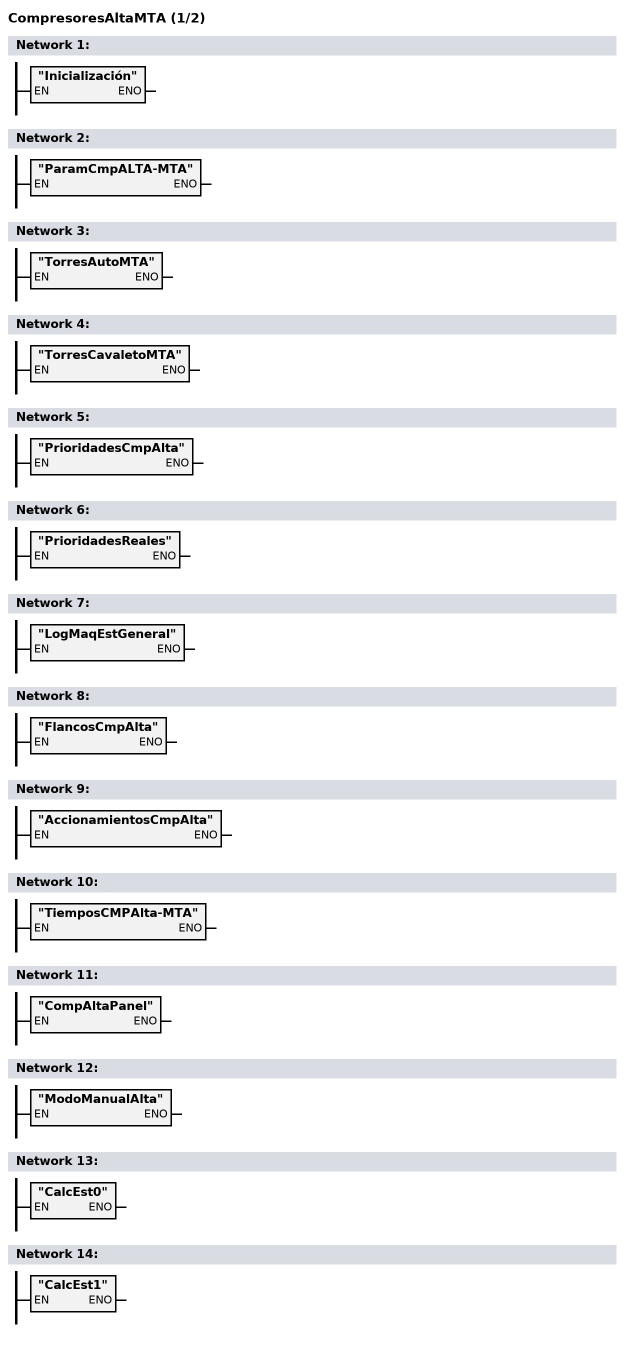
   RUNG wire#powerrail
      "Inicialización"()
   END_RUNG
   // the same network as SCL:
   "Inicialización"();
END_REGION

REGION Network 2
   RUNG wire#powerrail
      "ParamCmpALTA-MTA"()
   END_RUNG
   // the same network as SCL:
   "ParamCmpALTA-MTA"();
END_REGION

REGION Network 3
   RUNG wire#powerrail
      "TorresAutoMTA"()
   END_RUNG
   // the same network as SCL:
   "TorresAutoMTA"();
END_REGION

REGION Network 4
   RUNG wire#powerrail
      "TorresCavaletoMTA"()
   END_RUNG
   // the same network as SCL:
   "TorresCavaletoMTA"();
END_REGION

REGION Network 5
   RUNG wire#powerrail
      "PrioridadesCmpAlta"()
   END_RUNG
   // the same network as SCL:
   "PrioridadesCmpAlta"();
END_REGION

REGION Network 6
   RUNG wire#powerrail
      "PrioridadesReales"()
   END_RUNG
   // the same network as SCL:
   "PrioridadesReales"();
END_REGION

REGION Network 7
   RUNG wire#powerrail
      "LogMaqEstGeneral"()
   END_RUNG
   // the same network as SCL:
   "LogMaqEstGeneral"();
END_REGION

REGION Network 8
   RUNG wire#powerrail
      "FlancosCmpAlta"()
   END_RUNG
   // the same network as SCL:
   "FlancosCmpAlta"();
END_REGION

REGION Network 9
   RUNG wire#powerrail
      "AccionamientosCmpAlta"()
   END_RUNG
   // the same network as SCL:
   "AccionamientosCmpAlta"();
END_REGION

REGION Network 10
   RUNG wire#powerrail
      "TiemposCMPAlta-MTA"()
   END_RUNG
   // the same network as SCL:
   "TiemposCMPAlta-MTA"();
END_REGION

REGION Network 11
   RUNG wire#powerrail
      "CompAltaPanel"()
   END_RUNG
   // the same network as SCL:
   "CompAltaPanel"();
END_REGION

REGION Network 12
   RUNG wire#powerrail
      "ModoManualAlta"()
   END_RUNG
   // the same network as SCL:
   "ModoManualAlta"();
END_REGION

REGION Network 13
   RUNG wire#powerrail
      "CalcEst0"()
   END_RUNG
   // the same network as SCL:
   "CalcEst0"();
END_REGION

REGION Network 14
   RUNG wire#powerrail
      "CalcEst1"()
   END_RUNG
   // the same network as SCL:
   "CalcEst1"();
END_REGION

REGION Network 15
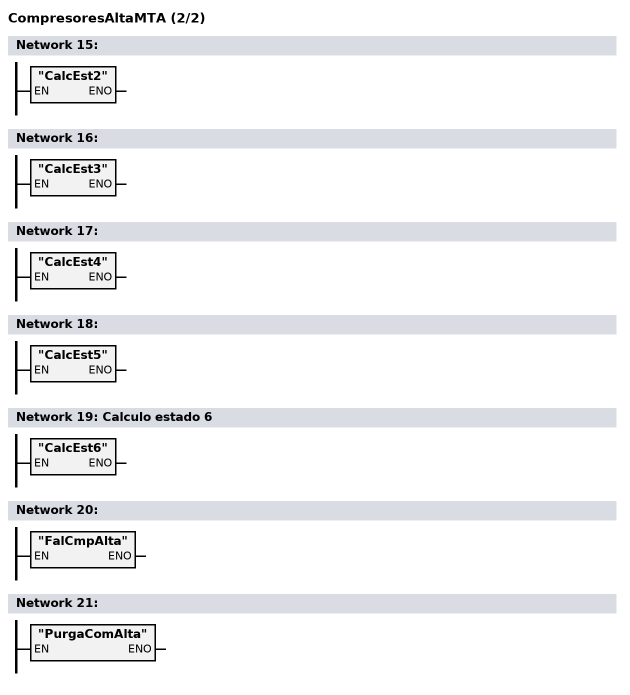
   RUNG wire#powerrail
      "CalcEst2"()
   END_RUNG
   // the same network as SCL:
   "CalcEst2"();
END_REGION

REGION Network 16
   RUNG wire#powerrail
      "CalcEst3"()
   END_RUNG
   // the same network as SCL:
   "CalcEst3"();
END_REGION

REGION Network 17
   RUNG wire#powerrail
      "CalcEst4"()
   END_RUNG
   // the same network as SCL:
   "CalcEst4"();
END_REGION

REGION Network 18
   RUNG wire#powerrail
      "CalcEst5"()
   END_RUNG
   // the same network as SCL:
   "CalcEst5"();
END_REGION

REGION Network 19: Calculo estado 6
   RUNG wire#powerrail
      "CalcEst6"()
   END_RUNG
   // the same network as SCL:
   "CalcEst6"();
END_REGION

REGION Network 20
   RUNG wire#powerrail
      "FalCmpAlta"()
   END_RUNG
   // the same network as SCL:
   "FalCmpAlta"();
END_REGION

REGION Network 21
   RUNG wire#powerrail
      "PurgaComAlta"()
   END_RUNG
   // the same network as SCL:
   "PurgaComAlta"();
END_REGION
END_FUNCTION

FUNCTION "ParamCmpALTA-MTA" : Void   // FC30, LAD
{ S7_Optimized_Access := 'FALSE' }
VERSION : 0.1
BEGIN

REGION Network 1
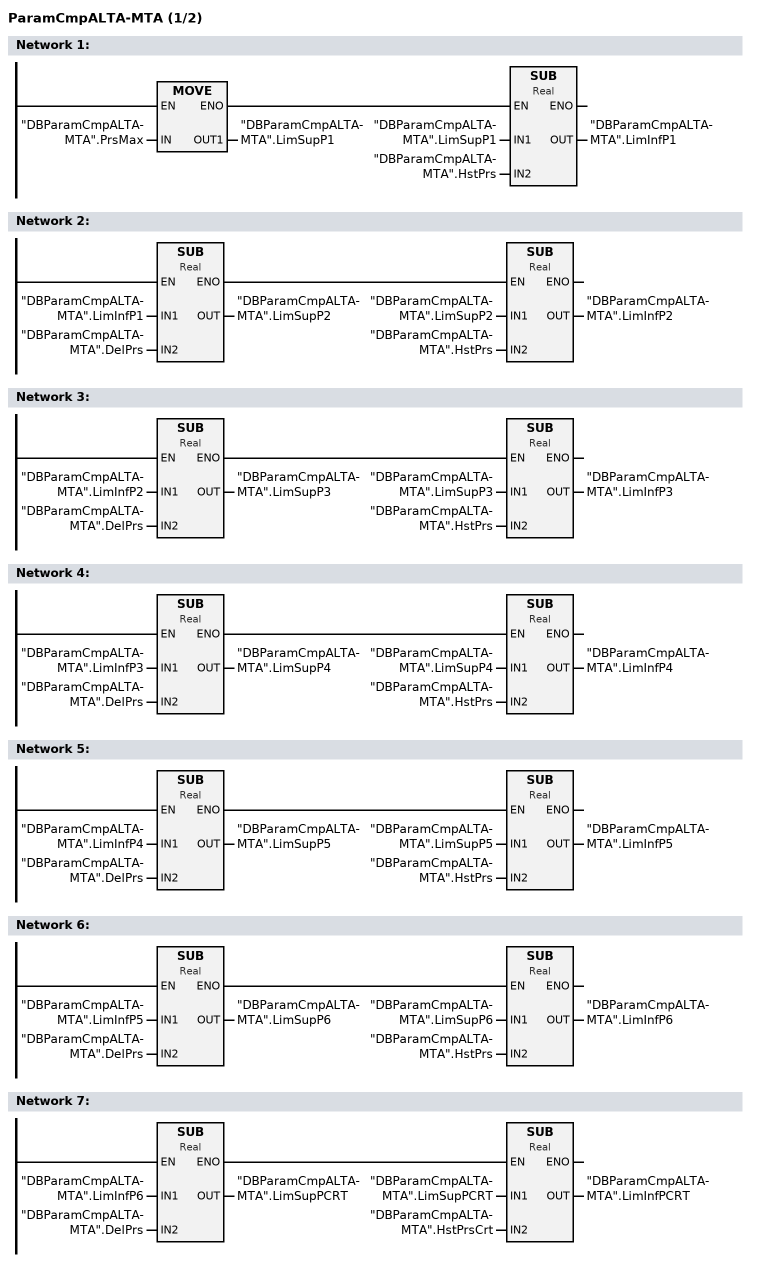
   RUNG wire#powerrail
      { S7_GenerateENO := "TRUE" } Move(in := "DBParamCmpALTA-MTA".PrsMax, out1 => "DBParamCmpALTA-MTA".LimSupP1)
      { S7_Templates := "SrcType := Real"; S7_GenerateENO := "TRUE" } Sub(in1 := "DBParamCmpALTA-MTA".LimSupP1, in2 := "DBParamCmpALTA-MTA".HstPrs, out => "DBParamCmpALTA-MTA".LimInfP1)
   END_RUNG
   // the same network as SCL:
   // ENO of a box is taken as its EN; it also drops when the box reports an error
   "DBParamCmpALTA-MTA".LimSupP1 := "DBParamCmpALTA-MTA".PrsMax;
   "DBParamCmpALTA-MTA".LimInfP1 := "DBParamCmpALTA-MTA".LimSupP1 - "DBParamCmpALTA-MTA".HstPrs;
END_REGION

REGION Network 2
   RUNG wire#powerrail
      { S7_Templates := "SrcType := Real"; S7_GenerateENO := "TRUE" } Sub(in1 := "DBParamCmpALTA-MTA".LimInfP1, in2 := "DBParamCmpALTA-MTA".DelPrs, out => "DBParamCmpALTA-MTA".LimSupP2)
      { S7_Templates := "SrcType := Real"; S7_GenerateENO := "TRUE" } Sub(in1 := "DBParamCmpALTA-MTA".LimSupP2, in2 := "DBParamCmpALTA-MTA".HstPrs, out => "DBParamCmpALTA-MTA".LimInfP2)
   END_RUNG
   // the same network as SCL:
   // ENO of a box is taken as its EN; it also drops when the box reports an error
   "DBParamCmpALTA-MTA".LimSupP2 := "DBParamCmpALTA-MTA".LimInfP1 - "DBParamCmpALTA-MTA".DelPrs;
   "DBParamCmpALTA-MTA".LimInfP2 := "DBParamCmpALTA-MTA".LimSupP2 - "DBParamCmpALTA-MTA".HstPrs;
END_REGION

REGION Network 3
   RUNG wire#powerrail
      { S7_Templates := "SrcType := Real"; S7_GenerateENO := "TRUE" } Sub(in1 := "DBParamCmpALTA-MTA".LimInfP2, in2 := "DBParamCmpALTA-MTA".DelPrs, out => "DBParamCmpALTA-MTA".LimSupP3)
      { S7_Templates := "SrcType := Real"; S7_GenerateENO := "TRUE" } Sub(in1 := "DBParamCmpALTA-MTA".LimSupP3, in2 := "DBParamCmpALTA-MTA".HstPrs, out => "DBParamCmpALTA-MTA".LimInfP3)
   END_RUNG
   // the same network as SCL:
   // ENO of a box is taken as its EN; it also drops when the box reports an error
   "DBParamCmpALTA-MTA".LimSupP3 := "DBParamCmpALTA-MTA".LimInfP2 - "DBParamCmpALTA-MTA".DelPrs;
   "DBParamCmpALTA-MTA".LimInfP3 := "DBParamCmpALTA-MTA".LimSupP3 - "DBParamCmpALTA-MTA".HstPrs;
END_REGION

REGION Network 4
   RUNG wire#powerrail
      { S7_Templates := "SrcType := Real"; S7_GenerateENO := "TRUE" } Sub(in1 := "DBParamCmpALTA-MTA".LimInfP3, in2 := "DBParamCmpALTA-MTA".DelPrs, out => "DBParamCmpALTA-MTA".LimSupP4)
      { S7_Templates := "SrcType := Real"; S7_GenerateENO := "TRUE" } Sub(in1 := "DBParamCmpALTA-MTA".LimSupP4, in2 := "DBParamCmpALTA-MTA".HstPrs, out => "DBParamCmpALTA-MTA".LimInfP4)
   END_RUNG
   // the same network as SCL:
   // ENO of a box is taken as its EN; it also drops when the box reports an error
   "DBParamCmpALTA-MTA".LimSupP4 := "DBParamCmpALTA-MTA".LimInfP3 - "DBParamCmpALTA-MTA".DelPrs;
   "DBParamCmpALTA-MTA".LimInfP4 := "DBParamCmpALTA-MTA".LimSupP4 - "DBParamCmpALTA-MTA".HstPrs;
END_REGION

REGION Network 5
   RUNG wire#powerrail
      { S7_Templates := "SrcType := Real"; S7_GenerateENO := "TRUE" } Sub(in1 := "DBParamCmpALTA-MTA".LimInfP4, in2 := "DBParamCmpALTA-MTA".DelPrs, out => "DBParamCmpALTA-MTA".LimSupP5)
      { S7_Templates := "SrcType := Real"; S7_GenerateENO := "TRUE" } Sub(in1 := "DBParamCmpALTA-MTA".LimSupP5, in2 := "DBParamCmpALTA-MTA".HstPrs, out => "DBParamCmpALTA-MTA".LimInfP5)
   END_RUNG
   // the same network as SCL:
   // ENO of a box is taken as its EN; it also drops when the box reports an error
   "DBParamCmpALTA-MTA".LimSupP5 := "DBParamCmpALTA-MTA".LimInfP4 - "DBParamCmpALTA-MTA".DelPrs;
   "DBParamCmpALTA-MTA".LimInfP5 := "DBParamCmpALTA-MTA".LimSupP5 - "DBParamCmpALTA-MTA".HstPrs;
END_REGION

REGION Network 6
   RUNG wire#powerrail
      { S7_Templates := "SrcType := Real"; S7_GenerateENO := "TRUE" } Sub(in1 := "DBParamCmpALTA-MTA".LimInfP5, in2 := "DBParamCmpALTA-MTA".DelPrs, out => "DBParamCmpALTA-MTA".LimSupP6)
      { S7_Templates := "SrcType := Real"; S7_GenerateENO := "TRUE" } Sub(in1 := "DBParamCmpALTA-MTA".LimSupP6, in2 := "DBParamCmpALTA-MTA".HstPrs, out => "DBParamCmpALTA-MTA".LimInfP6)
   END_RUNG
   // the same network as SCL:
   // ENO of a box is taken as its EN; it also drops when the box reports an error
   "DBParamCmpALTA-MTA".LimSupP6 := "DBParamCmpALTA-MTA".LimInfP5 - "DBParamCmpALTA-MTA".DelPrs;
   "DBParamCmpALTA-MTA".LimInfP6 := "DBParamCmpALTA-MTA".LimSupP6 - "DBParamCmpALTA-MTA".HstPrs;
END_REGION

REGION Network 7
   RUNG wire#powerrail
      { S7_Templates := "SrcType := Real"; S7_GenerateENO := "TRUE" } Sub(in1 := "DBParamCmpALTA-MTA".LimInfP6, in2 := "DBParamCmpALTA-MTA".DelPrs, out => "DBParamCmpALTA-MTA".LimSupPCRT)
      { S7_Templates := "SrcType := Real"; S7_GenerateENO := "TRUE" } Sub(in1 := "DBParamCmpALTA-MTA".LimSupPCRT, in2 := "DBParamCmpALTA-MTA".HstPrsCrt, out => "DBParamCmpALTA-MTA".LimInfPCRT)
   END_RUNG
   // the same network as SCL:
   // ENO of a box is taken as its EN; it also drops when the box reports an error
   "DBParamCmpALTA-MTA".LimSupPCRT := "DBParamCmpALTA-MTA".LimInfP6 - "DBParamCmpALTA-MTA".DelPrs;
   "DBParamCmpALTA-MTA".LimInfPCRT := "DBParamCmpALTA-MTA".LimSupPCRT - "DBParamCmpALTA-MTA".HstPrsCrt;
END_REGION

REGION Network 8: Falla General Flujostato Cavaleto
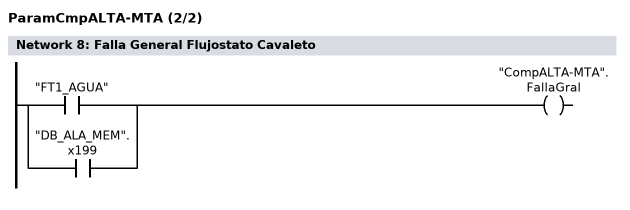
   RUNG wire#powerrail
      Contact( "FT1_AGUA" )
      wire#w1
      Coil( "CompALTA-MTA".FallaGral )
   END_RUNG
   RUNG wire#powerrail
      Contact( "DB_ALA_MEM".x199 )
   END_RUNG wire#w1
   // the same network as SCL:
   "CompALTA-MTA".FallaGral := "FT1_AGUA" OR "DB_ALA_MEM".x199;
END_REGION
END_FUNCTION

FUNCTION "TiemposCMPAlta-MTA" : Void   // FC31, LAD
{ S7_Optimized_Access := 'FALSE' }
VERSION : 0.1
   VAR_TEMP
      TEMP0 : Int;
   END_VAR
   VAR_TEMP   // added for the SCL form of the ladder/FBD networks
      _s5time1 : S5Time;
   END_VAR
BEGIN

REGION Network 1
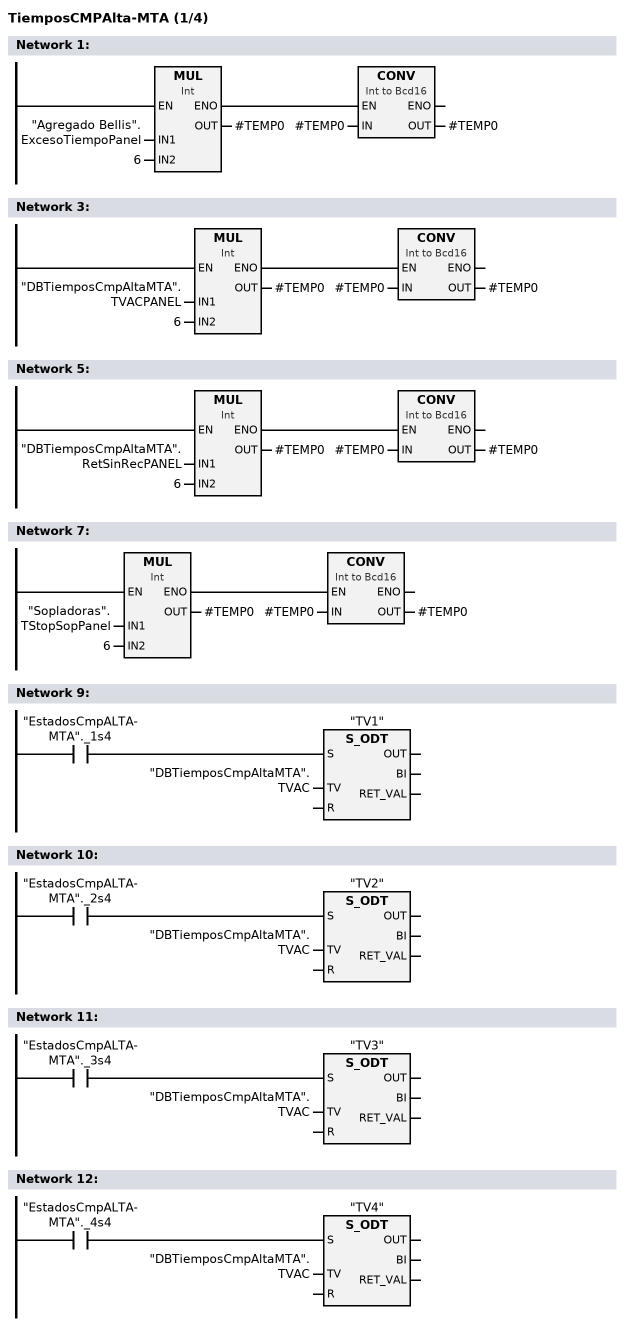
   RUNG wire#powerrail
      { S7_Templates := "SrcType := Int"; S7_GenerateENO := "TRUE" } Mul(in1 := "Agregado Bellis".ExcesoTiempoPanel, in2 := 6, out => #TEMP0)
      { S7_Templates := "[SrcType := Int, DestType := Bcd16]"; S7_GenerateENO := "TRUE" } Convert(in := #TEMP0, out => #TEMP0)
   END_RUNG
   // the same network as SCL:
   // ENO of a box is taken as its EN; it also drops when the box reports an error
   #TEMP0 := "Agregado Bellis".ExcesoTiempoPanel * 6;
   #TEMP0 := INT_TO_BCD16(#TEMP0);
END_REGION

REGION Network 2 (STL)
         L     12288;
         L     #TEMP0;
         OW;
         T     "Agregado Bellis".ExcesoTiempo;
         NOP   0;
END_REGION

REGION Network 3
   RUNG wire#powerrail
      { S7_Templates := "SrcType := Int"; S7_GenerateENO := "TRUE" } Mul(in1 := "DBTiemposCmpAltaMTA".TVACPANEL, in2 := 6, out => #TEMP0)
      { S7_Templates := "[SrcType := Int, DestType := Bcd16]"; S7_GenerateENO := "TRUE" } Convert(in := #TEMP0, out => #TEMP0)
   END_RUNG
   // the same network as SCL:
   // ENO of a box is taken as its EN; it also drops when the box reports an error
   #TEMP0 := "DBTiemposCmpAltaMTA".TVACPANEL * 6;
   #TEMP0 := INT_TO_BCD16(#TEMP0);
END_REGION

REGION Network 4 (STL)
         L     12288;
         L     #TEMP0;
         OW;
         T     "DBTiemposCmpAltaMTA".TVAC;
         NOP   0;
END_REGION

REGION Network 5
   RUNG wire#powerrail
      { S7_Templates := "SrcType := Int"; S7_GenerateENO := "TRUE" } Mul(in1 := "DBTiemposCmpAltaMTA".RetSinRecPANEL, in2 := 6, out => #TEMP0)
      { S7_Templates := "[SrcType := Int, DestType := Bcd16]"; S7_GenerateENO := "TRUE" } Convert(in := #TEMP0, out => #TEMP0)
   END_RUNG
   // the same network as SCL:
   // ENO of a box is taken as its EN; it also drops when the box reports an error
   #TEMP0 := "DBTiemposCmpAltaMTA".RetSinRecPANEL * 6;
   #TEMP0 := INT_TO_BCD16(#TEMP0);
END_REGION

REGION Network 6 (STL)
         L     12288;
         L     #TEMP0;
         OW;
         T     "DBTiemposCmpAltaMTA".RetSinRec;
         NOP   0;
END_REGION

REGION Network 7
   RUNG wire#powerrail
      { S7_Templates := "SrcType := Int"; S7_GenerateENO := "TRUE" } Mul(in1 := "Sopladoras".TStopSopPanel, in2 := 6, out => #TEMP0)
      { S7_Templates := "[SrcType := Int, DestType := Bcd16]"; S7_GenerateENO := "TRUE" } Convert(in := #TEMP0, out => #TEMP0)
   END_RUNG
   // the same network as SCL:
   // ENO of a box is taken as its EN; it also drops when the box reports an error
   #TEMP0 := "Sopladoras".TStopSopPanel * 6;
   #TEMP0 := INT_TO_BCD16(#TEMP0);
END_REGION

REGION Network 8 (STL)
         L     12288;
         L     #TEMP0;
         OW;
         T     "Sopladoras".TStopSop;
         NOP   0;
END_REGION

REGION Network 9
   RUNG wire#powerrail
      Contact( "EstadosCmpALTA-MTA"._1s4 )
      S_ODT(T_NO := "TV1", TV := "DBTiemposCmpAltaMTA".TVAC, R :=, BI =>, RET_VAL =>)
   END_RUNG
   // the same network as SCL:
   #_s5time1 := S_ODT(T_NO := "TV1", S := "EstadosCmpALTA-MTA"._1s4, TV := "DBTiemposCmpAltaMTA".TVAC);
END_REGION

REGION Network 10
   RUNG wire#powerrail
      Contact( "EstadosCmpALTA-MTA"._2s4 )
      S_ODT(T_NO := "TV2", TV := "DBTiemposCmpAltaMTA".TVAC, R :=, BI =>, RET_VAL =>)
   END_RUNG
   // the same network as SCL:
   #_s5time1 := S_ODT(T_NO := "TV2", S := "EstadosCmpALTA-MTA"._2s4, TV := "DBTiemposCmpAltaMTA".TVAC);
END_REGION

REGION Network 11
   RUNG wire#powerrail
      Contact( "EstadosCmpALTA-MTA"._3s4 )
      S_ODT(T_NO := "TV3", TV := "DBTiemposCmpAltaMTA".TVAC, R :=, BI =>, RET_VAL =>)
   END_RUNG
   // the same network as SCL:
   #_s5time1 := S_ODT(T_NO := "TV3", S := "EstadosCmpALTA-MTA"._3s4, TV := "DBTiemposCmpAltaMTA".TVAC);
END_REGION

REGION Network 12
   RUNG wire#powerrail
      Contact( "EstadosCmpALTA-MTA"._4s4 )
      S_ODT(T_NO := "TV4", TV := "DBTiemposCmpAltaMTA".TVAC, R :=, BI =>, RET_VAL =>)
   END_RUNG
   // the same network as SCL:
   #_s5time1 := S_ODT(T_NO := "TV4", S := "EstadosCmpALTA-MTA"._4s4, TV := "DBTiemposCmpAltaMTA".TVAC);
END_REGION

REGION Network 13
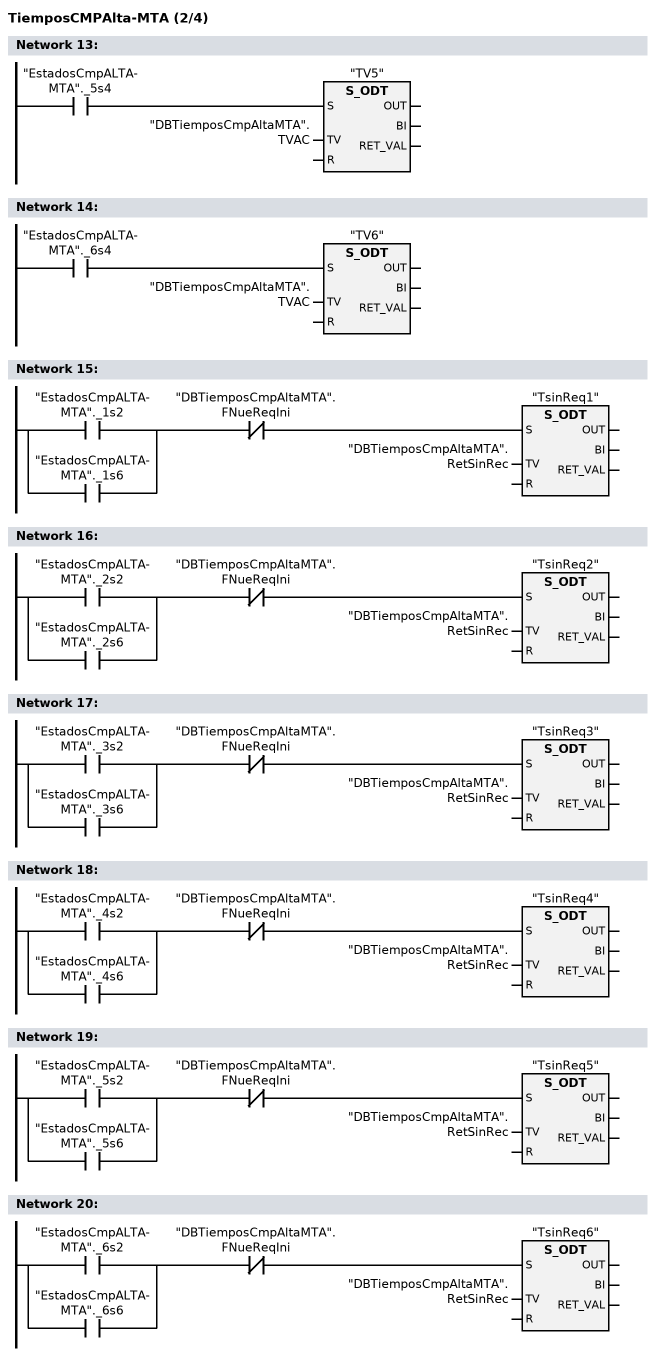
   RUNG wire#powerrail
      Contact( "EstadosCmpALTA-MTA"._5s4 )
      S_ODT(T_NO := "TV5", TV := "DBTiemposCmpAltaMTA".TVAC, R :=, BI =>, RET_VAL =>)
   END_RUNG
   // the same network as SCL:
   #_s5time1 := S_ODT(T_NO := "TV5", S := "EstadosCmpALTA-MTA"._5s4, TV := "DBTiemposCmpAltaMTA".TVAC);
END_REGION

REGION Network 14
   RUNG wire#powerrail
      Contact( "EstadosCmpALTA-MTA"._6s4 )
      S_ODT(T_NO := "TV6", TV := "DBTiemposCmpAltaMTA".TVAC, R :=, BI =>, RET_VAL =>)
   END_RUNG
   // the same network as SCL:
   #_s5time1 := S_ODT(T_NO := "TV6", S := "EstadosCmpALTA-MTA"._6s4, TV := "DBTiemposCmpAltaMTA".TVAC);
END_REGION

REGION Network 15
   RUNG wire#powerrail
      Contact( "EstadosCmpALTA-MTA"._1s2 )
      wire#w1
      I_Contact( "DBTiemposCmpAltaMTA".FNueReqIni )
      S_ODT(T_NO := "TsinReq1", TV := "DBTiemposCmpAltaMTA".RetSinRec, R :=, BI =>, RET_VAL =>)
   END_RUNG
   RUNG wire#powerrail
      Contact( "EstadosCmpALTA-MTA"._1s6 )
   END_RUNG wire#w1
   // the same network as SCL:
   #_s5time1 := S_ODT(T_NO := "TsinReq1",
                      S := ("EstadosCmpALTA-MTA"._1s2 OR "EstadosCmpALTA-MTA"._1s6) AND NOT "DBTiemposCmpAltaMTA".FNueReqIni,
                      TV := "DBTiemposCmpAltaMTA".RetSinRec);
END_REGION

REGION Network 16
   RUNG wire#powerrail
      Contact( "EstadosCmpALTA-MTA"._2s2 )
      wire#w1
      I_Contact( "DBTiemposCmpAltaMTA".FNueReqIni )
      S_ODT(T_NO := "TsinReq2", TV := "DBTiemposCmpAltaMTA".RetSinRec, R :=, BI =>, RET_VAL =>)
   END_RUNG
   RUNG wire#powerrail
      Contact( "EstadosCmpALTA-MTA"._2s6 )
   END_RUNG wire#w1
   // the same network as SCL:
   #_s5time1 := S_ODT(T_NO := "TsinReq2",
                      S := ("EstadosCmpALTA-MTA"._2s2 OR "EstadosCmpALTA-MTA"._2s6) AND NOT "DBTiemposCmpAltaMTA".FNueReqIni,
                      TV := "DBTiemposCmpAltaMTA".RetSinRec);
END_REGION

REGION Network 17
   RUNG wire#powerrail
      Contact( "EstadosCmpALTA-MTA"._3s2 )
      wire#w1
      I_Contact( "DBTiemposCmpAltaMTA".FNueReqIni )
      S_ODT(T_NO := "TsinReq3", TV := "DBTiemposCmpAltaMTA".RetSinRec, R :=, BI =>, RET_VAL =>)
   END_RUNG
   RUNG wire#powerrail
      Contact( "EstadosCmpALTA-MTA"._3s6 )
   END_RUNG wire#w1
   // the same network as SCL:
   #_s5time1 := S_ODT(T_NO := "TsinReq3",
                      S := ("EstadosCmpALTA-MTA"._3s2 OR "EstadosCmpALTA-MTA"._3s6) AND NOT "DBTiemposCmpAltaMTA".FNueReqIni,
                      TV := "DBTiemposCmpAltaMTA".RetSinRec);
END_REGION

REGION Network 18
   RUNG wire#powerrail
      Contact( "EstadosCmpALTA-MTA"._4s2 )
      wire#w1
      I_Contact( "DBTiemposCmpAltaMTA".FNueReqIni )
      S_ODT(T_NO := "TsinReq4", TV := "DBTiemposCmpAltaMTA".RetSinRec, R :=, BI =>, RET_VAL =>)
   END_RUNG
   RUNG wire#powerrail
      Contact( "EstadosCmpALTA-MTA"._4s6 )
   END_RUNG wire#w1
   // the same network as SCL:
   #_s5time1 := S_ODT(T_NO := "TsinReq4",
                      S := ("EstadosCmpALTA-MTA"._4s2 OR "EstadosCmpALTA-MTA"._4s6) AND NOT "DBTiemposCmpAltaMTA".FNueReqIni,
                      TV := "DBTiemposCmpAltaMTA".RetSinRec);
END_REGION

REGION Network 19
   RUNG wire#powerrail
      Contact( "EstadosCmpALTA-MTA"._5s2 )
      wire#w1
      I_Contact( "DBTiemposCmpAltaMTA".FNueReqIni )
      S_ODT(T_NO := "TsinReq5", TV := "DBTiemposCmpAltaMTA".RetSinRec, R :=, BI =>, RET_VAL =>)
   END_RUNG
   RUNG wire#powerrail
      Contact( "EstadosCmpALTA-MTA"._5s6 )
   END_RUNG wire#w1
   // the same network as SCL:
   #_s5time1 := S_ODT(T_NO := "TsinReq5",
                      S := ("EstadosCmpALTA-MTA"._5s2 OR "EstadosCmpALTA-MTA"._5s6) AND NOT "DBTiemposCmpAltaMTA".FNueReqIni,
                      TV := "DBTiemposCmpAltaMTA".RetSinRec);
END_REGION

REGION Network 20
   RUNG wire#powerrail
      Contact( "EstadosCmpALTA-MTA"._6s2 )
      wire#w1
      I_Contact( "DBTiemposCmpAltaMTA".FNueReqIni )
      S_ODT(T_NO := "TsinReq6", TV := "DBTiemposCmpAltaMTA".RetSinRec, R :=, BI =>, RET_VAL =>)
   END_RUNG
   RUNG wire#powerrail
      Contact( "EstadosCmpALTA-MTA"._6s6 )
   END_RUNG wire#w1
   // the same network as SCL:
   #_s5time1 := S_ODT(T_NO := "TsinReq6",
                      S := ("EstadosCmpALTA-MTA"._6s2 OR "EstadosCmpALTA-MTA"._6s6) AND NOT "DBTiemposCmpAltaMTA".FNueReqIni,
                      TV := "DBTiemposCmpAltaMTA".RetSinRec);
END_REGION

REGION Network 21
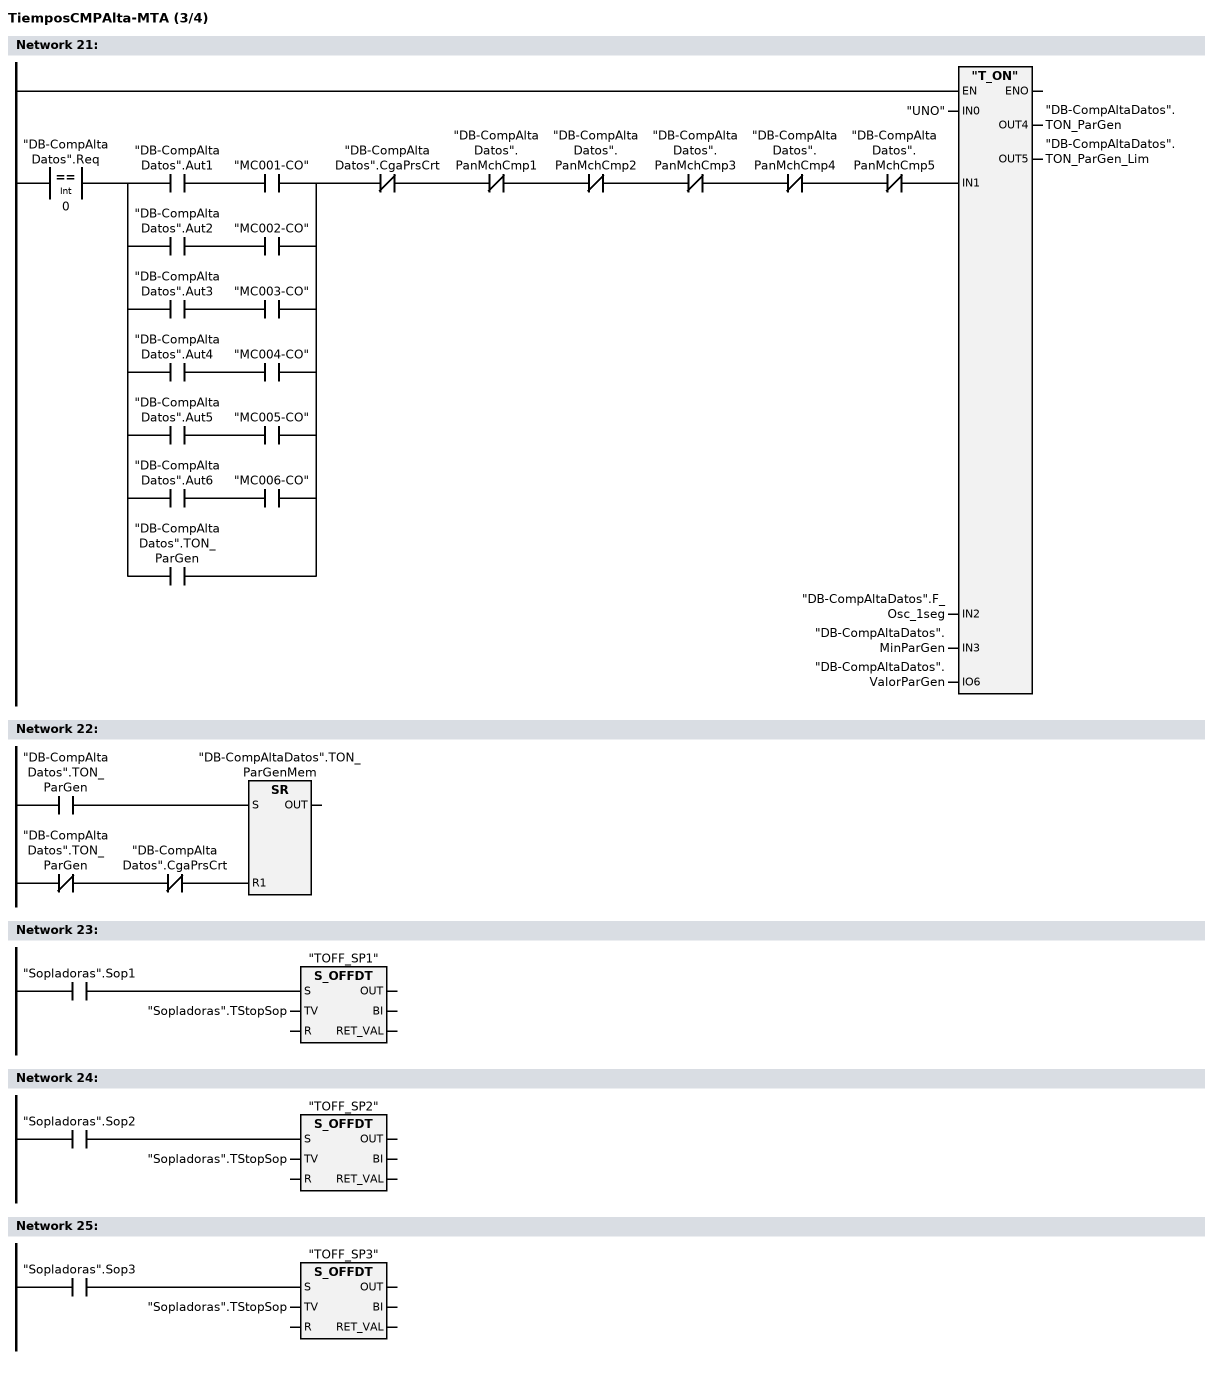
   RUNG wire#powerrail
      "T_ON"(IN1 := wire#w3, IN0 := "UNO", IN2 := "DB-CompAltaDatos".F_Osc_1seg, IN3 := "DB-CompAltaDatos".MinParGen, IO6 := "DB-CompAltaDatos".ValorParGen, OUT4 => "DB-CompAltaDatos".TON_ParGen, OUT5 => "DB-CompAltaDatos".TON_ParGen_Lim)
   END_RUNG
   RUNG wire#powerrail
      { S7_Templates := "SrcType := Int" } EQ_Contact(in1 := "DB-CompAltaDatos".Req, in2 := 0)
      wire#w1
      Contact( "DB-CompAltaDatos".Aut1 )
      Contact( "MC001-CO" )
      wire#w2
      I_Contact( "DB-CompAltaDatos".CgaPrsCrt )
      I_Contact( "DB-CompAltaDatos".PanMchCmp1 )
      I_Contact( "DB-CompAltaDatos".PanMchCmp2 )
      I_Contact( "DB-CompAltaDatos".PanMchCmp3 )
      I_Contact( "DB-CompAltaDatos".PanMchCmp4 )
      I_Contact( "DB-CompAltaDatos".PanMchCmp5 )
   END_RUNG wire#w3
   RUNG wire#w1
      Contact( "DB-CompAltaDatos".Aut2 )
      Contact( "MC002-CO" )
   END_RUNG wire#w2
   RUNG wire#w1
      Contact( "DB-CompAltaDatos".Aut3 )
      Contact( "MC003-CO" )
   END_RUNG wire#w2
   RUNG wire#w1
      Contact( "DB-CompAltaDatos".Aut4 )
      Contact( "MC004-CO" )
   END_RUNG wire#w2
   RUNG wire#w1
      Contact( "DB-CompAltaDatos".Aut5 )
      Contact( "MC005-CO" )
   END_RUNG wire#w2
   RUNG wire#w1
      Contact( "DB-CompAltaDatos".Aut6 )
      Contact( "MC006-CO" )
   END_RUNG wire#w2
   RUNG wire#w1
      Contact( "DB-CompAltaDatos".TON_ParGen )
   END_RUNG wire#w2
   // the same network as SCL:
   "T_ON"(IN0 := "UNO",
          IN1 := ("DB-CompAltaDatos".Req = 0) AND (("DB-CompAltaDatos".Aut1 AND "MC001-CO") OR ("DB-CompAltaDatos".Aut2 AND "MC002-CO") OR ("DB-CompAltaDatos".Aut3 AND "MC003-CO") OR ("DB-CompAltaDatos".Aut4 AND "MC004-CO") OR ("DB-CompAltaDatos".Aut5 AND "MC005-CO") OR ("DB-CompAltaDatos".Aut6 AND "MC006-CO") OR "DB-CompAltaDatos".TON_ParGen) AND NOT "DB-CompAltaDatos".CgaPrsCrt AND NOT "DB-CompAltaDatos".PanMchCmp1 AND NOT "DB-CompAltaDatos".PanMchCmp2 AND NOT "DB-CompAltaDatos".PanMchCmp3 AND NOT "DB-CompAltaDatos".PanMchCmp4 AND NOT "DB-CompAltaDatos".PanMchCmp5,
          IN2 := "DB-CompAltaDatos".F_Osc_1seg,
          IN3 := "DB-CompAltaDatos".MinParGen,
          IO6 := "DB-CompAltaDatos".ValorParGen,
          OUT4 => "DB-CompAltaDatos".TON_ParGen,
          OUT5 => "DB-CompAltaDatos".TON_ParGen_Lim);
END_REGION

REGION Network 22
   RUNG wire#powerrail
      Contact( "DB-CompAltaDatos".TON_ParGen )
      S_SR(operand := "DB-CompAltaDatos".TON_ParGenMem, r1 := wire#w1)
   END_RUNG
   RUNG wire#powerrail
      I_Contact( "DB-CompAltaDatos".TON_ParGen )
      I_Contact( "DB-CompAltaDatos".CgaPrsCrt )
   END_RUNG wire#w1
   // the same network as SCL:
   IF "DB-CompAltaDatos".TON_ParGen THEN
       "DB-CompAltaDatos".TON_ParGenMem := TRUE;   // SR flip-flop
   END_IF;
   IF NOT "DB-CompAltaDatos".TON_ParGen AND NOT "DB-CompAltaDatos".CgaPrsCrt THEN
       "DB-CompAltaDatos".TON_ParGenMem := FALSE;
   END_IF;
END_REGION

REGION Network 23
   RUNG wire#powerrail
      Contact( "Sopladoras".Sop1 )
      S_OFFDT(T_NO := "TOFF_SP1", TV := "Sopladoras".TStopSop, R :=, BI =>, RET_VAL =>)
   END_RUNG
   // the same network as SCL:
   #_s5time1 := S_OFFDT(T_NO := "TOFF_SP1", TV := "Sopladoras".TStopSop, S := "Sopladoras".Sop1);
END_REGION

REGION Network 24
   RUNG wire#powerrail
      Contact( "Sopladoras".Sop2 )
      S_OFFDT(T_NO := "TOFF_SP2", TV := "Sopladoras".TStopSop, R :=, BI =>, RET_VAL =>)
   END_RUNG
   // the same network as SCL:
   #_s5time1 := S_OFFDT(T_NO := "TOFF_SP2", TV := "Sopladoras".TStopSop, S := "Sopladoras".Sop2);
END_REGION

REGION Network 25
   RUNG wire#powerrail
      Contact( "Sopladoras".Sop3 )
      S_OFFDT(T_NO := "TOFF_SP3", TV := "Sopladoras".TStopSop, R :=, BI =>, RET_VAL =>)
   END_RUNG
   // the same network as SCL:
   #_s5time1 := S_OFFDT(T_NO := "TOFF_SP3", TV := "Sopladoras".TStopSop, S := "Sopladoras".Sop3);
END_REGION

REGION Network 26
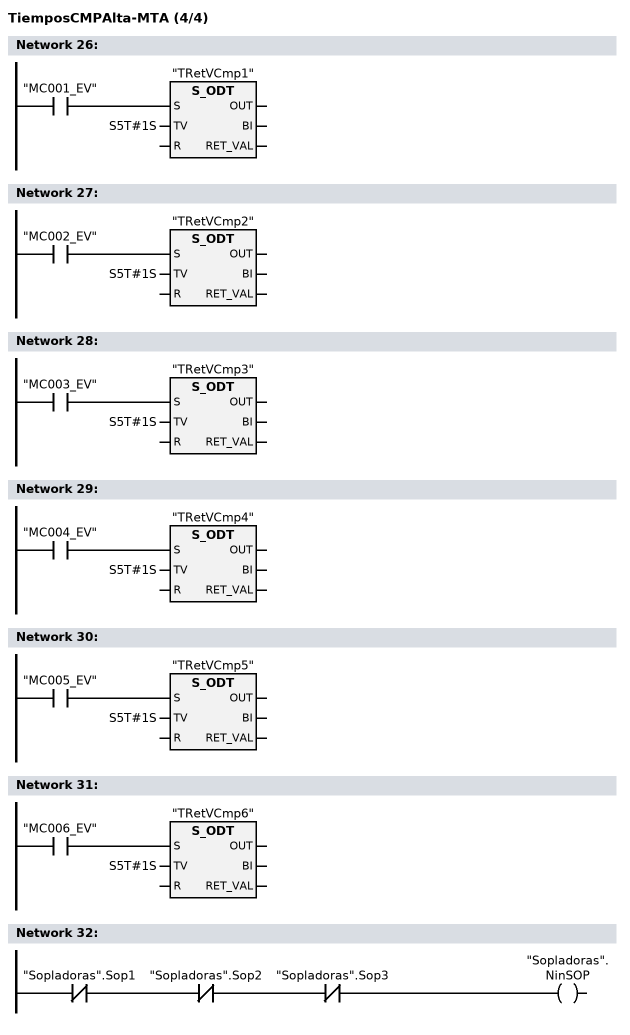
   RUNG wire#powerrail
      Contact( "MC001_EV" )
      S_ODT(T_NO := "TRetVCmp1", TV := S5T#1S, R :=, BI =>, RET_VAL =>)
   END_RUNG
   // the same network as SCL:
   #_s5time1 := S_ODT(T_NO := "TRetVCmp1", TV := S5T#1S, S := "MC001_EV");
END_REGION

REGION Network 27
   RUNG wire#powerrail
      Contact( "MC002_EV" )
      S_ODT(T_NO := "TRetVCmp2", TV := S5T#1S, R :=, BI =>, RET_VAL =>)
   END_RUNG
   // the same network as SCL:
   #_s5time1 := S_ODT(T_NO := "TRetVCmp2", TV := S5T#1S, S := "MC002_EV");
END_REGION

REGION Network 28
   RUNG wire#powerrail
      Contact( "MC003_EV" )
      S_ODT(T_NO := "TRetVCmp3", TV := S5T#1S, R :=, BI =>, RET_VAL =>)
   END_RUNG
   // the same network as SCL:
   #_s5time1 := S_ODT(T_NO := "TRetVCmp3", TV := S5T#1S, S := "MC003_EV");
END_REGION

REGION Network 29
   RUNG wire#powerrail
      Contact( "MC004_EV" )
      S_ODT(T_NO := "TRetVCmp4", TV := S5T#1S, R :=, BI =>, RET_VAL =>)
   END_RUNG
   // the same network as SCL:
   #_s5time1 := S_ODT(T_NO := "TRetVCmp4", TV := S5T#1S, S := "MC004_EV");
END_REGION

REGION Network 30
   RUNG wire#powerrail
      Contact( "MC005_EV" )
      S_ODT(T_NO := "TRetVCmp5", TV := S5T#1S, R :=, BI =>, RET_VAL =>)
   END_RUNG
   // the same network as SCL:
   #_s5time1 := S_ODT(T_NO := "TRetVCmp5", TV := S5T#1S, S := "MC005_EV");
END_REGION

REGION Network 31
   RUNG wire#powerrail
      Contact( "MC006_EV" )
      S_ODT(T_NO := "TRetVCmp6", TV := S5T#1S, R :=, BI =>, RET_VAL =>)
   END_RUNG
   // the same network as SCL:
   #_s5time1 := S_ODT(T_NO := "TRetVCmp6", S := "MC006_EV", TV := S5T#1S);
END_REGION

REGION Network 32
   RUNG wire#powerrail
      I_Contact( "Sopladoras".Sop1 )
      I_Contact( "Sopladoras".Sop2 )
      I_Contact( "Sopladoras".Sop3 )
      Coil( "Sopladoras".NinSOP )
   END_RUNG
   // the same network as SCL:
   "Sopladoras".NinSOP := NOT "Sopladoras".Sop1 AND NOT "Sopladoras".Sop2 AND NOT "Sopladoras".Sop3;
END_REGION
END_FUNCTION

FUNCTION "T_ON" : Void   // FC32, LAD
{ S7_Optimized_Access := 'FALSE' }
VERSION : 0.1
   VAR_INPUT
      IN0 : Bool;
      IN1 : Bool;
      IN2 : Bool;
      IN3 : Int;
   END_VAR
   VAR_OUTPUT
      OUT4 : Bool;
      OUT5 : Bool;
   END_VAR
   VAR_IN_OUT
      IO6 : Int;
   END_VAR
   VAR_TEMP
      TEMP7 : Int;
      TEMP8 : Int;
   END_VAR
   VAR_TEMP   // added for the SCL form of the ladder/FBD networks
      _w1 : Bool;
   END_VAR
BEGIN

REGION Network 1
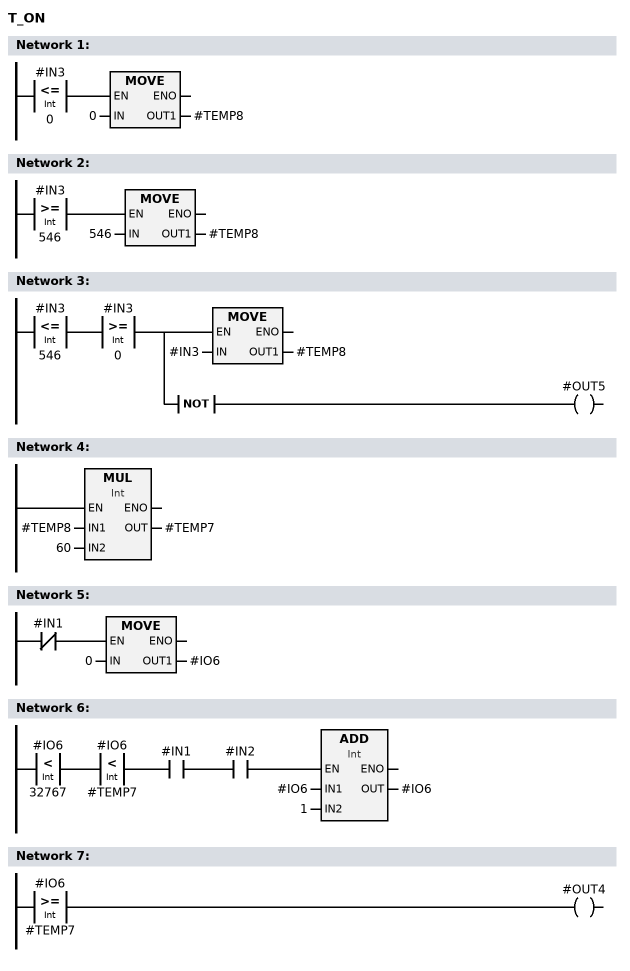
   RUNG wire#powerrail
      { S7_Templates := "SrcType := Int" } LE_Contact(in1 := #IN3, in2 := 0)
      { S7_GenerateENO := "TRUE" } Move(in := 0, out1 => #TEMP8)
   END_RUNG
   // the same network as SCL:
   IF #IN3 <= 0 THEN #TEMP8 := 0; END_IF;
END_REGION

REGION Network 2
   RUNG wire#powerrail
      { S7_Templates := "SrcType := Int" } GE_Contact(in1 := #IN3, in2 := 546)
      { S7_GenerateENO := "TRUE" } Move(in := 546, out1 => #TEMP8)
   END_RUNG
   // the same network as SCL:
   IF #IN3 >= 546 THEN #TEMP8 := 546; END_IF;
END_REGION

REGION Network 3
   RUNG wire#powerrail
      { S7_Templates := "SrcType := Int" } LE_Contact(in1 := #IN3, in2 := 546)
      { S7_Templates := "SrcType := Int" } GE_Contact(in1 := #IN3, in2 := 0)
      wire#w1
      { S7_GenerateENO := "TRUE" } Move(in := #IN3, out1 => #TEMP8)
   END_RUNG
   RUNG wire#w1
      Not()
      Coil( #OUT5 )
   END_RUNG
   // the same network as SCL:
   #_w1 := (#IN3 <= 546) AND (#IN3 >= 0);
   IF #_w1 THEN #TEMP8 := #IN3; END_IF;
   #OUT5 := NOT #_w1;
END_REGION

REGION Network 4
   RUNG wire#powerrail
      { S7_Templates := "SrcType := Int"; S7_GenerateENO := "TRUE" } Mul(in1 := #TEMP8, in2 := 60, out => #TEMP7)
   END_RUNG
   // the same network as SCL:
   #TEMP7 := #TEMP8 * 60;
END_REGION

REGION Network 5
   RUNG wire#powerrail
      I_Contact( #IN1 )
      { S7_GenerateENO := "TRUE" } Move(in := 0, out1 => #IO6)
   END_RUNG
   // the same network as SCL:
   IF NOT #IN1 THEN #IO6 := 0; END_IF;
END_REGION

REGION Network 6
   RUNG wire#powerrail
      { S7_Templates := "SrcType := Int" } LT_Contact(in1 := #IO6, in2 := 32767)
      { S7_Templates := "SrcType := Int" } LT_Contact(in1 := #IO6, in2 := #TEMP7)
      Contact( #IN1 )
      Contact( #IN2 )
      { S7_Templates := "SrcType := Int"; S7_GenerateENO := "TRUE" } Add(in1 := #IO6, in2 := 1, out => #IO6)
   END_RUNG
   // the same network as SCL:
   IF (#IO6 < 32767) AND (#IO6 < #TEMP7) AND #IN1 AND #IN2 THEN #IO6 := #IO6 + 1; END_IF;
END_REGION

REGION Network 7
   RUNG wire#powerrail
      { S7_Templates := "SrcType := Int" } GE_Contact(in1 := #IO6, in2 := #TEMP7)
      Coil( #OUT4 )
   END_RUNG
   // the same network as SCL:
   #OUT4 := #IO6 >= #TEMP7;
END_REGION
END_FUNCTION

FUNCTION "PrioridadesCmpAlta" : Void   // FC33, LAD
{ S7_Optimized_Access := 'FALSE' }
VERSION : 0.1
   VAR_TEMP   // added for the SCL form of the ladder/FBD networks
      _w1 : Bool;
   END_VAR
BEGIN

REGION Network 1